// TIA Portal project "IntercambioDeDatos" (V16)

(* hardware
DEVICE "PC-System"  CPU 1515SP PC
   slot 0: "PC-System"  CPU 1515SP PC F  6ES7 677-2SBx2-0xB0  V20.8
      slot 124: "Diagbase"  Diagbase  V6.0.4
      slot 125: "PC-System"  PC Station 2.7  Station_Manager  V2.7
   slot 2: "PROFINET onboard_2"  IE General  IE_CP  V2.2.0
      slot 1: "Puerto_1"  X2 P1
   slot 3: "Software PLC_1"  CPU 1505SP F  6ES7 672-5SC11-0YA0  V2.7
      slot 3: "Display de la CPU_1"  6ES7591-1BA00-0AA0
   slot 127: "BA 2xRJ45"  BA 2xRJ45  6ES7 193-6AR00-0AA0  V0.0
      slot 32769: "Puerto_1"  X1 P1  6ES7 193-6AR00-0AA0
      slot 32770: "Puerto_2"  X1 P2  6ES7 193-6AR00-0AA0
   slot 1006: "Módulo servidor_1"  Server module  6ES7 193-6PA00-0AA0  V1.1
      slot 1: "Módulo servidor_1"  Server module
DEVICE "Dispositivo GSD_1"  GSD.Device.PN
   slot 0: "Rack"  Rack  V1.0
   slot 0: "URIODev1"  V1.0  00000
      slot 0: "V1.0"  V1.0
      slot 1: "Interface"  Interface
         slot 1: "RJ45 10/100 MBit/s"  RJ45 10/100 MBit/s
   slot 1: "1_T2O State_1"  1_T2O State  1.0
      slot 0: "1_T2O State"  1_T2O State
   slot 2: "2_T2O IO_1"  2_T2O IO  1.0
      slot 0: "2_T2O IO"  2_T2O IO
   slot 3: "3_T2O Joints_1"  3_T2O Joints  1.0
      slot 0: "3_T2O Joints"  3_T2O Joints
   slot 4: "4_T2O TCP_1"  4_T2O TCP  1.0
      slot 0: "4_T2O TCP"  4_T2O TCP
   slot 5: "5_T2O General Purpose Bit Registers_1"  5_T2O General Purpose Bit Registers  1.0
      slot 0: "5_T2O General Purpose Bit Registers"  5_T2O General Purpose Bit Registers
   slot 6: "6_T2O General Purpose Int Registers_1"  6_T2O General Purpose Int Registers  1.0
      slot 0: "6_T2O General Purpose Int Registers"  6_T2O General Purpose Int Registers
   slot 7: "7_T2O General Purpose Float Registers_1"  7_T2O General Purpose Float Registers  1.0
      slot 0: "7_T2O General Purpose Float Registers"  7_T2O General Purpose Float Registers
   slot 8: "8_O2T Robot IO_1"  8_O2T Robot IO  1.0
      slot 0: "8_O2T Robot IO"  8_O2T Robot IO
   slot 9: "9_O2T General Purpose Registers 1_1"  9_O2T General Purpose Registers 1  1.0
      slot 0: "9_O2T General Purpose Registers 1"  9_O2T General Purpose Registers 1
   slot 10: "10_O2T General Purpose Registers 2_1"  10_O2T General Purpose Registers 2  1.0
      slot 0: "10_O2T General Purpose Registers 2"  10_O2T General Purpose Registers 2
DEVICE "HMI"  KTP1200 Basic PN
   slot 0: "HMI_2"  KTP1200 Basic PN  6AV2 123-2MB03-0AX0  16.0.0.0
   slot 1: "HMI_RT_1"  KTP1200 Basic PN  6AV2 123-2MB03-0AX0  16.0.0.0
   slot 5: "HMI_2.IE_CP_1"  PROFINET Interface  16.0.0.0
      slot 1: "Interfaz PROFINET_1"  PROFINET Interface
         slot 1: "Port_1"  Port
*)

// ===== PLC "Software PLC_1"  CPU 1505SP F =====

VAR_GLOBAL   // PLC tag table "Tabla de variables estándar"
   "Flanco_Marcha" AT %M0.4 : Bool;
   "Biestable_Marcha" AT %M10.0 : Bool;
   "Tag_2" AT %M11.0 : Bool;
   "Tag_1" AT %MW20 : Int;
   "Tag_3" AT %MW22 : Int;
   "Tag_4" AT %MW24 : Int;
END_VAR

VAR_GLOBAL   // PLC tag table "IntercambioDeDatos_Variables"
   "URI" AT %I0.0 : "UR_T2O";   // Grupo de variables en donde se guardan los valores que se envian al robot
   "URO" AT %Q0.0 : "UR_O2T";   // Grupo de variables en donde se guardan los valores que llegan desde el robot
   "Marcha" AT %M0.0 : Bool;   // Variable que define en que momento debe comenzar funcionar el robot
   "Servicio_Completado" AT %M0.1 : Bool;
   "Servicio" AT %MW3 : Int;   // Variable que define el número de servicio a ejecutar
   "CantPiezas" AT %MW5 : Int;   // Variable que define la cantidad de pieza que se deben realizar.
   "Aux" AT %M1.7 : Bool;
   "No_Item_Completados" AT %MW7 : Int;
   "Item_Completado" AT %M0.2 : Bool;
   "Marcha_Reset" AT %M0.3 : Bool;
   "Flag_New_Service" AT %M0.5 : Bool;
   "MqttConnected" AT %M1.0 : Bool;
   "MqttDataReceived" AT %M1.1 : Bool;
   "Serialize" AT %M1.2 : Bool;
   "MqttSubscribed" AT %M1.3 : Bool;
   "MqttPreviousStatus" AT %MW9 : Word;
   "MqttUnsuscribed" AT %M1.4 : Bool;
   "Marcha_aux" AT %M0.6 : Bool;
   "Flanco_Service_Compl" AT %M0.7 : Bool;
   "Aux_Initial_Time_Stamp" AT %M12.0 : ULInt;
   "Aux_Final_Time_Stamp" AT %M20.0 : ULInt;
   "Aux_Service_Time_Stamp" AT %M28.0 : ULInt;
END_VAR

// folder: Common

TYPE "typeDiagnostics"
TITLE = typeDiagnostics
// Provides a structure for detailed diagnostics
   STRUCT
      status : Word;   // Status of the block or error identification when error occurred
      subfunctionStatus : DWord;   // Status or return value of called FBs, FCs and system blocks
      stateNumber : DInt;   // State in the state machine of the block where the error occurred
   END_STRUCT;
END_TYPE

// folder: LMQTT

TYPE "LMQTT_typeConnParams"
TITLE = LMQTT_typeConnParams
// Specifies connection parameters for the mqtt connection
   STRUCT
      hwId : Hw_Any;   // Hardware identifier of the interface. 0: interface is selected automatically
      connId : Conn_Ouc;   // Unique connection identifier
      brokerAddress : Struct   // Information on the MQTT broker
         qdnAddress : String;   // Fully qualified domain name of the broker. must end with a dot "."
         ipAddress : IP_V4;   // If no FQDN is used, enter ip-address of the broker instead
         port : UInt;   // Enter the port of the mqtt broker
      END_STRUCT;
      tls : Struct   // Parameters for TLS encryption
         enableTls : Bool;   // TRUE: Enables TLS, FALSE: disable TLS
         validateServerIdentity : Bool;   // TRUE: Validate server certificate, FALSE: No validation of server certificate
         brokerCert : UDInt;   // ID of the broker's certificate in TIA Portal
         clientCert : UDInt;   // ID of the client's certificate in TIA Portal
      END_STRUCT;
      keepAlive : UInt;   // Keepalive mechanism for MQTT in seconds. 0: disabled.
   END_STRUCT;
END_TYPE

// folder: LStream/DataTypes

TYPE "LStream_typeElement"
TITLE = LStream_typeElement
// describes the element for LStream libraries, by providing key-value pair and the depth of the element
   STRUCT
      "type" : SInt := -1;   // Type of element XML/JSON; -1 = inital value; 0 = Element/Object; 1 = Attribute/Array; 2 = Text/String; 3 = Number; 4 = Boolean / Type of element; -1 = inital value; 0 = Element/Object; 1 = Attribute/Array; 2 = Text
      key : String;   // Key name of element
      value : String := 'NULL';   // Value of element, null key has no value
      depth : SInt := -1;   // Depth of the key nesting
   END_STRUCT;
END_TYPE

// folder: Robot

TYPE "UR__O2T_Robot"
VERSION : 0.1
   STRUCT
      "SSM: Speed slider fraction mask" : Bool;
      Reserved_1 : Bool;
      Reserved_2 : Bool;
      Reserved_3 : Bool;
      Reserved_4 : Bool;
      Reserved_5 : Bool;
      Reserved_6 : Bool;
      Reserved_7 : Bool;
      Reserved_8_15 : USInt;
      Reserved_16_31 : UInt;
      "Speed slider fraction" : Real;
   END_STRUCT;
END_TYPE

TYPE "UR__O2T_ints"
VERSION : 0.1
   STRUCT
      Register : Array[0..11] of DInt;
   END_STRUCT;
END_TYPE

TYPE "UR__O2T_floats"
VERSION : 0.1
   STRUCT
      Register : Array[0..11] of Real;
   END_STRUCT;
END_TYPE

TYPE "UR__O2T_IOs"
VERSION : 0.1
   STRUCT
      "Standard digital output mask" : USInt;
      "Configurable digital output mask" : USInt;
      "Standard digital outputs" : USInt;
      "Configurable digital outputs" : USInt;
      "AOM: Analog output mask" : USInt;
      "AOT: Analog output types" : USInt;
      "TDOM: Tool digital output mask" : USInt;
      "TDO: Tool digital output" : USInt;
      "Standard analog output" : Array[0..1] of Real;
   END_STRUCT;
END_TYPE

TYPE "UR__O2T_bits"
VERSION : 0.1
   STRUCT
      Register : Array[0..31] of Bool;
   END_STRUCT;
END_TYPE

TYPE "UR_9_O2T_Registers"
VERSION : 0.1
   STRUCT
      Bits : "UR__O2T_bits";
      Ints : "UR__O2T_ints";
      Floats : "UR__O2T_floats";
   END_STRUCT;
END_TYPE

TYPE "UR_8_O2T_Robot_IO"
VERSION : 0.1
   STRUCT
      Robot : "UR__O2T_Robot";
      IOs : "UR__O2T_IOs";
   END_STRUCT;
END_TYPE

TYPE "UR__T2O_Safety"
VERSION : 0.1
   STRUCT
      "Safety mode" : USInt;
      Reserved_1 : USInt;
      Reserved_2 : UInt;
      "NO: Is normal mode" : Bool;
      "RD: Is reduced mode" : Bool;
      "PS: Is protective stopped" : Bool;
      "RC: Is recovery mode" : Bool;
      "SS: Is safeguard stopped" : Bool;
      "SES: Is system emergency stopped" : Bool;
      "RES: Is robot emergency stopped" : Bool;
      "ES: Is emergency stopped" : Bool;
      "VL: Is violation" : Bool;
      "FT: Is fault" : Bool;
      "ST: Is stopped due to safety" : Bool;
      Reserved_11 : Bool;
      Reserved_12 : Bool;
      Reserved_13 : Bool;
      Reserved_14 : Bool;
      Reserved_15 : Bool;
      Reserved_16_31 : UInt;
   END_STRUCT;
END_TYPE

TYPE "UR__T2O_Robot"
VERSION : 0.1
   STRUCT
      "Controller major version" : USInt;
      "Controller minor version" : USInt;
      Reserved : UInt;
      "Robot mode" : USInt;
      "Real time machine seconds" : USInt;
      "Real time machine milliseconds" : UInt;
      "Real time machine minutes" : USInt;
      "Real time machine hours" : USInt;
      "Real time machine days" : UInt;
      "Robot current [A]" : Real;
      "PW: Is power on" : Bool;
      "PR: Is program running" : Bool;
      "TB: Is teach button pressed" : Bool;
      "PB: Is power button pressed" : Bool;
      Reserved_4 : Bool;
      Reserved_5 : Bool;
      Reserved_6 : Bool;
      Reserved_7 : Bool;
      Reserved_8_15 : USInt;
      Reserved_16_31 : UInt;
      "Speed slider fraction" : Real;
   END_STRUCT;
END_TYPE

TYPE "UR__T2O_Tool"
VERSION : 0.1
   STRUCT
      "Tool mode" : USInt;
      Reserved_7_15 : USInt;
      Reserved_16_31 : UInt;
      "TDI: Tool Digital Inputs" : USInt;
      "TDO: Tool Digital Outputs" : USInt;
      "TAIT: Tool Analog Input Types" : USInt;
      Reserved_24_31 : USInt;
      "Tool analog input [A or V]" : Array[0..1] of Real;
      "Tool output voltage [V]" : Real;
      "Tool current [A]" : Real;
   END_STRUCT;
END_TYPE

TYPE "UR_O2T"
VERSION : 0.1
   STRUCT
      "Robot IO" : "UR_8_O2T_Robot_IO";
      "Reg 1" : "UR_9_O2T_Registers";
      "Reg 2" : "UR_9_O2T_Registers";
   END_STRUCT;
END_TYPE

TYPE "UR_4_T2O_TCP"
VERSION : 0.1
   STRUCT
      "TCP Position (X,Y,Z) [m]" : Array[0..2] of Real;
      "TCP Position (RX,RY,RZ) [rad]" : Array[0..2] of Real;
      "TCP velocity (X,Y,Z) [m/s]" : Array[0..2] of Real;
      "TCP velocity (RX,RY,RZ) [rad/s]" : Array[0..2] of Real;
      "TCP force (X,Y,Z) [N]" : Array[0..2] of Real;
      "TCP torque (X,Y,Z) [Nm]" : Array[0..2] of Real;
      "TCP force scalar [N]" : Real;
   END_STRUCT;
END_TYPE

TYPE "UR_3_T2O_Joints"
VERSION : 0.1
   STRUCT
      "Joint position [rad]" : Array[0..5] of Real;
      "Joint velocity [rad/s]" : Array[0..5] of Real;
      "Joint current [A]" : Array[0..5] of Real;
      "Joint temperature [°C]" : Array[0..5] of Real;
      "Joint mode" : Array[0..5] of USInt;
      Reserved_9 : UInt;
   END_STRUCT;
END_TYPE

TYPE "UR_2_T2O_IO"
VERSION : 0.1
   STRUCT
      IOs : "UR__T2O_IOs";
      Tool : "UR__T2O_Tool";
   END_STRUCT;
END_TYPE

TYPE "UR_1_T2O_State"
VERSION : 0.1
   STRUCT
      Robot : "UR__T2O_Robot";
      Safety : "UR__T2O_Safety";
   END_STRUCT;
END_TYPE

TYPE "UR_7_T2O_FloatRegisters"
VERSION : 0.1
   STRUCT
      Register : Array[0..23] of Real;
   END_STRUCT;
END_TYPE

TYPE "UR_6_T2O_IntRegisters"
VERSION : 0.1
   STRUCT
      Register : Array[0..23] of DInt;
   END_STRUCT;
END_TYPE

TYPE "UR_T2O"
VERSION : 0.1
   STRUCT
      State : "UR_1_T2O_State";
      IO : "UR_2_T2O_IO";
      Joints : "UR_3_T2O_Joints";
      TCP : "UR_4_T2O_TCP";
      Bits : "UR_5_T2O_BitRegisters";
      Ints : "UR_6_T2O_IntRegisters";
      Floats : "UR_7_T2O_FloatRegisters";
   END_STRUCT;
END_TYPE

TYPE "UR__T2O_IOs"
VERSION : 0.1
   STRUCT
      "Standard digital inputs" : USInt;
      "Configurable digital inputs" : USInt;
      "Standard digital outputs" : USInt;
      "Configurable digital outputs" : USInt;
      "Analog I/O types" : USInt;
      Reserved_8_15 : USInt;
      Reserved_16_31 : UInt;
      "Standard analog input [A or V]" : Array[0..1] of Real;
      "Standard analog output [A or V]" : Array[0..1] of Real;
      "I/O current [A]" : Real;
      "Euromap67 input bits" : Array[0..31] of Bool;
      "Euromap67 output bits" : Array[0..31] of Bool;
      "Euromap67 24V voltage" : Real;
      "Euromap67 24V current" : Real;
   END_STRUCT;
END_TYPE

TYPE "UR_5_T2O_BitRegisters"
VERSION : 0.1
   STRUCT
      Register : Array[0..63] of Bool;
   END_STRUCT;
END_TYPE

// folder: (top level)

DATA_BLOCK "Main_Safety_RTG1_DB"   // DB1, F_DB
{ S7_Optimized_Access := 'TRUE' }
NAME : FUSI
VERSION : 0.1
// stored: InstanceOfName Main_Safety_RTG1
"Main_Safety_RTG1"
BEGIN
END_DATA_BLOCK

DATA_BLOCK "MqttDB"   // DB3
{ S7_Optimized_Access := 'TRUE' }
AUTHOR : Siemens
FAMILY : LMQTT
VERSION : 1.0
   VAR
      control : Struct
         connect : Bool;
         publish : Bool;
         subscribe : Bool;
         unsubscribe : Bool;
      END_STRUCT;
      output : Struct
         valid : Bool;
         done : Bool;
         busy : Bool;
         error : Bool;
         status : Word;
         diagnostics : "typeDiagnostics";
      END_STRUCT;
      connparams : "LMQTT_typeConnParams";
      clientid : WString[20] := WSTRING#'Alazne';
      username : WString[20];
      password : WString[20];
      willtopic : WString[20] := WSTRING#'willTopic';
      willMessage : Array[0..99] of Byte;
      willmesscnt : UInt := 10;
      qos : USInt := 0;
      topic : WString[100] := WSTRING#'Operation';
      message : Array[0..999] of Byte;
      pubMessageCnt : UDInt := 1;
      retain : Bool;
      receivedTopic : WString[200];
      receivedmessage : Array[0..999] of Byte;
      receivedMsgLen : UDInt;
      receivedMsgStatus : USInt;
      dadoRecebido : String[100];
      dadoEnviado : String[100];
   END_VAR
BEGIN
   connparams.connId := 16#0001;
   connparams.brokerAddress.port := 1883;
   willMessage[0] := 16#6F;
   willMessage[1] := 16#66;
   willMessage[2] := 16#66;
   willMessage[3] := 16#6C;
   willMessage[4] := 16#69;
   willMessage[5] := 16#6E;
   willMessage[6] := 16#65;
   message[0] := 53;
   connparams.brokerAddress.ipAddress.ADDR[1] := 192;
   connparams.brokerAddress.ipAddress.ADDR[2] := 168;
   connparams.brokerAddress.ipAddress.ADDR[3] := 2;
   connparams.brokerAddress.ipAddress.ADDR[4] := 151;
   connparams.keepAlive := 30;   // Periodo de tiempo durante el cual se considera que una conexión esta viva sin que hay consexión entre el cliente y el bróker.
   connparams.hwId := 0;
END_DATA_BLOCK

DATA_BLOCK "AASassetDB"   // DB5
{ S7_Optimized_Access := 'TRUE' }
VERSION : 0.1
   VAR
      Control : Struct
         Flag_New_Service : Bool;
         Flag_Item_Completed : Bool;
         Flag_Service_Completed : Bool;
      END_STRUCT;
      Agent2PLC : Struct
         Id : Struct
            Machine_Reference : UDInt;
            Order_Reference : UDInt;
            Batch_Reference : UDInt;
            Ref_Subproduct_Type : UDInt;
         END_STRUCT;
         Operation : Struct
            Ref_Service_Type : UDInt;
            No_of_Items : USInt;
         END_STRUCT;
      END_STRUCT;
      PLC2Agent : Struct
         Id : Struct
            Machine_Reference : UDInt;
            Order_Reference : UDInt;
            Batch_Reference : UDInt;
            Ref_Subproduct_Type : UDInt;
            Ref_Service_Type : UDInt;
            Item_Number : USInt;
         END_STRUCT;
         Data : Struct
            Initial_Time_Stamp : LDT;
            Final_Time_Stamp : LDT;
            Service_Time_Stamp : LDT;
         END_STRUCT;
      END_STRUCT;
   END_VAR
BEGIN
END_DATA_BLOCK

DATA_BLOCK "JSON_DeserializParamDB"   // DB9
{ S7_Optimized_Access := 'TRUE' }
VERSION : 0.1
   VAR
      execute : Bool;
      search : Bool;
      jsonByteArray : Array[0..999] of Byte;
      tree : Array[0..999] of "LStream_typeElement";
      resultCount : Int;
      out : Struct
         done : Bool;
         busy : Bool;
         error : Bool;
         status : Word;
         resultCount : Int;
      END_STRUCT;
   END_VAR
BEGIN
END_DATA_BLOCK

DATA_BLOCK "JSON_SerializParamDB"   // DB10
{ S7_Optimized_Access := 'TRUE' }
VERSION : 0.1
   VAR
      execute : Bool;
      out : Struct
         done : Bool;
         busy : Bool;
         error : Bool;
         status : Word;
      END_STRUCT;
      tree : Array[0..999] of "LStream_typeElement";
      jsonByteArray : Array[0..999] of Byte;
      resultCount : Int;
   END_VAR
BEGIN
   tree[0]."type" := 0;
   tree[0].key := 'Control';
   tree[0].depth := 0;
   tree[1]."type" := 4;
   tree[1].key := 'Flag_Item_Completed';
   tree[1].depth := 1;
   tree[2]."type" := 4;
   tree[2].key := 'Flag_Service_Completed';
   tree[2].depth := 1;
   tree[3]."type" := 0;
   tree[3].key := 'Id';
   tree[3].depth := 0;
   tree[4]."type" := 3;
   tree[4].key := 'Machine_Reference';
   tree[4].depth := 1;
   tree[5]."type" := 3;
   tree[5].key := 'Order_Reference';
   tree[5].depth := 1;
   tree[6]."type" := 3;
   tree[6].key := 'Batch_Reference';
   tree[6].depth := 1;
   tree[7]."type" := 3;
   tree[7].key := 'Ref_Subproduct_Type';
   tree[7].depth := 1;
   tree[8].key := 'Ref_Service_Type';
   tree[8]."type" := 3;
   tree[8].depth := 1;
   tree[9]."type" := 3;
   tree[9].key := 'Item_Number';
   tree[9].depth := 1;
   tree[10]."type" := 0;
   tree[10].key := 'Data';
   tree[10].depth := 0;
   tree[11]."type" := 3;
   tree[11].key := 'Initial_Time_Stamp';
   tree[11].depth := 1;
   tree[12]."type" := 3;
   tree[12].key := 'Final_Time_Stamp';
   tree[12].depth := 1;
   tree[13]."type" := 3;
   tree[13].key := 'Service_Time_Stamp';
   tree[13].depth := 1;
END_DATA_BLOCK

// folder: LMQTT

DATA_BLOCK "LMQTT_Client_DB"   // DB2
{ S7_Optimized_Access := 'TRUE' }
AUTHOR : SUP
FAMILY : LMQTT
VERSION : 3.0
// stored: InstanceOfName LMQTT_Client
"LMQTT_Client"
BEGIN
END_DATA_BLOCK

// folder: LStream

DATA_BLOCK "LStream_JsonDeserializer_DB"   // DB7
{ S7_Optimized_Access := 'TRUE' }
AUTHOR : DI_FA_S_SUP_EuC
FAMILY : LStream
VERSION : 1.0
// stored: InstanceOfName LStream_JsonDeserializer
"LStream_JsonDeserializer"
BEGIN
END_DATA_BLOCK

DATA_BLOCK "LStream_JsonSerializer_DB"   // DB8
{ S7_Optimized_Access := 'TRUE' }
AUTHOR : DI_FA_S_SUP_EuC
FAMILY : LStream
VERSION : 1.0
// stored: InstanceOfName LStream_JsonSerializer
"LStream_JsonSerializer"
BEGIN
END_DATA_BLOCK

// folder: (top level)

FUNCTION_BLOCK "Main_Safety_RTG1"   // FB1, F_FBD
{ S7_Optimized_Access := 'TRUE' }
BEGIN
END_FUNCTION_BLOCK

FUNCTION "Outputs2LStreamTree" : Void   // FC1, SCL
{ S7_Optimized_Access := 'TRUE' }
VERSION : 0.1
BEGIN
   // Asignación de valores 
   (* "JSON_SerializParamDB".tree[1].value := "AASassetDb".Control.Flag_Item_Completed; *)

   (* "JSON_SerializParamDB".tree[1].value := 'false';
   "JSON_SerializParamDB".tree[2].value := 'false'; *)
   (* "JSON_SerializParamDB".tree[4].value := '123';
   "JSON_SerializParamDB".tree[5].value := '22';
   "JSON_SerializParamDB".tree[6].value := '33';
   "JSON_SerializParamDB".tree[7].value := '99'; *)

   IF "AASassetDB".Control.Flag_Service_Completed = 1 THEN
       "JSON_SerializParamDB".tree[2].value := 'true';
   ELSE
       "JSON_SerializParamDB".tree[2].value := 'false';
   END_IF;

   IF "AASassetDB".Control.Flag_Item_Completed = 1 THEN
       "JSON_SerializParamDB".tree[1].value := 'true';
   ELSE
       "JSON_SerializParamDB".tree[1].value := 'false';
   END_IF;

   "JSON_SerializParamDB".tree[4].value := UDINT_TO_STRING("AASassetDB".PLC2Agent.Id.Machine_Reference);
   "JSON_SerializParamDB".tree[5].value := UDINT_TO_STRING("AASassetDB".PLC2Agent.Id.Order_Reference);
   "JSON_SerializParamDB".tree[6].value := UDINT_TO_STRING("AASassetDB".PLC2Agent.Id.Batch_Reference);
   "JSON_SerializParamDB".tree[7].value := UDINT_TO_STRING("AASassetDB".PLC2Agent.Id.Ref_Subproduct_Type);
   "JSON_SerializParamDB".tree[8].value := UDINT_TO_STRING("AASassetDB".PLC2Agent.Id.Ref_Service_Type);
   "JSON_SerializParamDB".tree[9].value := USINT_TO_STRING("AASassetDB".PLC2Agent.Id.Item_Number);

   "JSON_SerializParamDB".tree[11].value := ULINT_TO_STRING(LDT_TO_ULINT("AASassetDB".PLC2Agent.Data.Initial_Time_Stamp));
   "JSON_SerializParamDB".tree[12].value := ULINT_TO_STRING(LDT_TO_ULINT("AASassetDB".PLC2Agent.Data.Final_Time_Stamp));
   "JSON_SerializParamDB".tree[13].value := ULINT_TO_STRING(LDT_TO_ULINT("AASassetDB".PLC2Agent.Data.Service_Time_Stamp));
END_FUNCTION

FUNCTION "LStreamTree2Inputs" : Void   // FC3, SCL
{ S7_Optimized_Access := 'TRUE' }
VERSION : 0.1
   VAR_TEMP
      Indice : Int;
   END_VAR
BEGIN
   // Volcado de los valores recibidos del bróker en las variables del DB.

   // Id
   "AASassetDB".Agent2PLC.Id.Machine_Reference := STRING_TO_UDINT("JSON_DeserializParamDB".tree[8].value);
   "AASassetDB".Agent2PLC.Id.Order_Reference := STRING_TO_UDINT("JSON_DeserializParamDB".tree[7].value);
   "AASassetDB".Agent2PLC.Id.Batch_Reference := STRING_TO_UDINT("JSON_DeserializParamDB".tree[5].value);
   "AASassetDB".Agent2PLC.Id.Ref_Subproduct_Type := STRING_TO_UDINT("JSON_DeserializParamDB".tree[6].value);

   // Operation
   "AASassetDB".Agent2PLC.Operation.Ref_Service_Type := STRING_TO_UDINT("JSON_DeserializParamDB".tree[11].value);
   "AASassetDB".Agent2PLC.Operation.No_of_Items := STRING_TO_USINT("JSON_DeserializParamDB".tree[10].value);
END_FUNCTION

ORGANIZATION_BLOCK "Main"   // OB1, LAD, ProgramCycle
TITLE = "Main Program Sweep (Cycle)"
{ S7_Optimized_Access := 'TRUE' }
VERSION : 0.1
   VAR_INPUT
      Initial_Call : Bool;   // Initial call of this OB
      Remanence : Bool;   // =True, if remanent data are available
   END_VAR
   VAR_TEMP
      FlancoNeg_Item_Completed : Bool;
      FlancoPos_Item_Completed : Bool;
   END_VAR
   VAR_TEMP   // added for the SCL form of the ladder/FBD networks
      _w1 : Bool;
      _w2 : Bool;
   END_VAR
BEGIN

REGION Network 1: Cliente MQTT
   // En este segmento nos encargamos tanto de la suscripción a un tópico como de las publicaciones que se realizarán en el tópico de publicaciones.
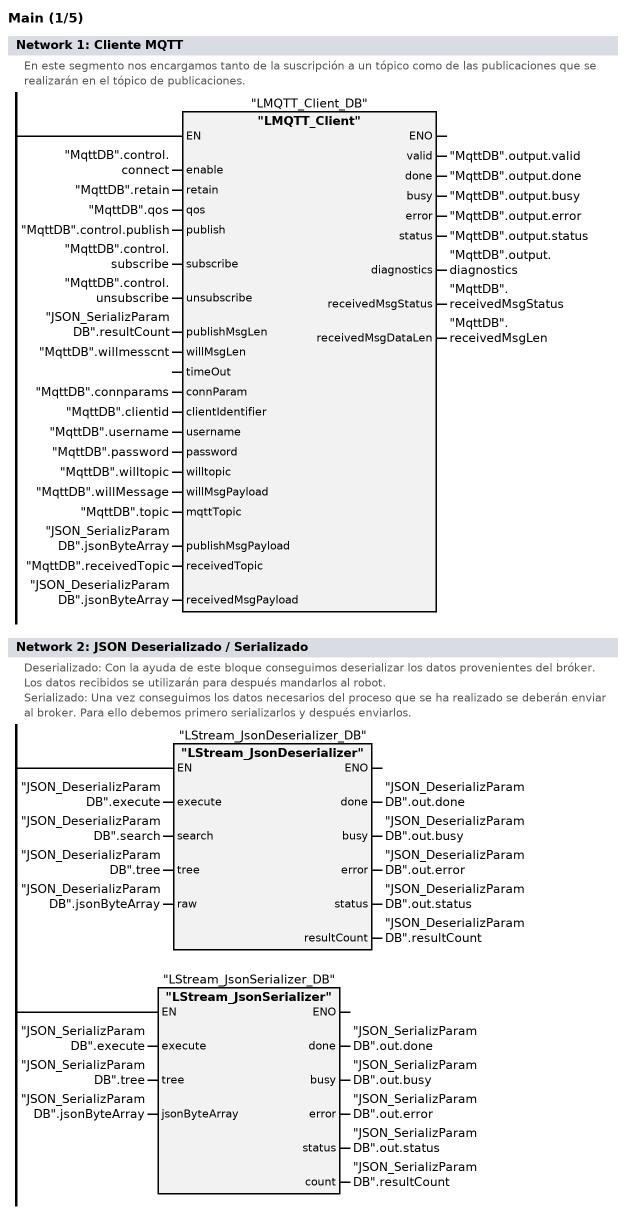
   RUNG wire#powerrail
      "LMQTT_Client_DB"(enable := "MqttDB".control.connect, retain := "MqttDB".retain, qos := "MqttDB".qos, publish := "MqttDB".control.publish, subscribe := "MqttDB".control.subscribe, unsubscribe := "MqttDB".control.unsubscribe, publishMsgLen := "JSON_SerializParamDB".resultCount, willMsgLen := "MqttDB".willmesscnt, timeOut :=, connParam := "MqttDB".connparams, clientIdentifier := "MqttDB".clientid, username := "MqttDB".username, password := "MqttDB".password, willtopic := "MqttDB".willtopic, willMsgPayload := "MqttDB".willMessage, mqttTopic := "MqttDB".topic, publishMsgPayload := "JSON_SerializParamDB".jsonByteArray, receivedTopic := "MqttDB".receivedTopic, receivedMsgPayload := "JSON_DeserializParamDB".jsonByteArray, valid => "MqttDB".output.valid, done => "MqttDB".output.done, busy => "MqttDB".output.busy, error => "MqttDB".output.error, status => "MqttDB".output.status, diagnostics => "MqttDB".output.diagnostics, receivedMsgStatus => "MqttDB".receivedMsgStatus, receivedMsgDataLen => "MqttDB".receivedMsgLen)
   END_RUNG
   // the same network as SCL:
   "LMQTT_Client_DB"(enable := "MqttDB".control.connect,   // "LMQTT_Client"
                     retain := "MqttDB".retain,
                     qos := "MqttDB".qos,
                     publish := "MqttDB".control.publish,
                     subscribe := "MqttDB".control.subscribe,
                     unsubscribe := "MqttDB".control.unsubscribe,
                     publishMsgLen := "JSON_SerializParamDB".resultCount,
                     willMsgLen := "MqttDB".willmesscnt,
                     connParam := "MqttDB".connparams,
                     clientIdentifier := "MqttDB".clientid,
                     username := "MqttDB".username,
                     password := "MqttDB".password,
                     willtopic := "MqttDB".willtopic,
                     willMsgPayload := "MqttDB".willMessage,
                     mqttTopic := "MqttDB".topic,
                     publishMsgPayload := "JSON_SerializParamDB".jsonByteArray,
                     receivedTopic := "MqttDB".receivedTopic,
                     receivedMsgPayload := "JSON_DeserializParamDB".jsonByteArray,
                     valid => "MqttDB".output.valid,
                     done => "MqttDB".output.done,
                     busy => "MqttDB".output.busy,
                     error => "MqttDB".output.error,
                     status => "MqttDB".output.status,
                     diagnostics => "MqttDB".output.diagnostics,
                     receivedMsgStatus => "MqttDB".receivedMsgStatus,
                     receivedMsgDataLen => "MqttDB".receivedMsgLen);
END_REGION

REGION Network 2: JSON Deserializado / Serializado
   // Deserializado: Con la ayuda de este bloque conseguimos deserializar los datos provenientes del bróker. 
   // Los datos recibidos se utilizarán para después mandarlos al robot.
   // 
   // Serializado: Una vez conseguimos los datos necesarios del proceso que se ha realizado se deberán enviar al broker. Para ello debemos primero serializarlos y después enviarlos.
   RUNG wire#powerrail
      "LStream_JsonDeserializer_DB"(execute := "JSON_DeserializParamDB".execute, search := "JSON_DeserializParamDB".search, tree := "JSON_DeserializParamDB".tree, raw := "JSON_DeserializParamDB".jsonByteArray, done => "JSON_DeserializParamDB".out.done, busy => "JSON_DeserializParamDB".out.busy, error => "JSON_DeserializParamDB".out.error, status => "JSON_DeserializParamDB".out.status, resultCount => "JSON_DeserializParamDB".resultCount)
   END_RUNG
   RUNG wire#powerrail
      "LStream_JsonSerializer_DB"(execute := "JSON_SerializParamDB".execute, tree := "JSON_SerializParamDB".tree, jsonByteArray := "JSON_SerializParamDB".jsonByteArray, done => "JSON_SerializParamDB".out.done, busy => "JSON_SerializParamDB".out.busy, error => "JSON_SerializParamDB".out.error, status => "JSON_SerializParamDB".out.status, count => "JSON_SerializParamDB".resultCount)
   END_RUNG
   // the same network as SCL:
   "LStream_JsonDeserializer_DB"(execute := "JSON_DeserializParamDB".execute,   // "LStream_JsonDeserializer"
                           search := "JSON_DeserializParamDB".search,
                           tree := "JSON_DeserializParamDB".tree,
                           raw := "JSON_DeserializParamDB".jsonByteArray,
                           done => "JSON_DeserializParamDB".out.done,
                           busy => "JSON_DeserializParamDB".out.busy,
                           error => "JSON_DeserializParamDB".out.error,
                           status => "JSON_DeserializParamDB".out.status,
                           resultCount => "JSON_DeserializParamDB".resultCount);
   "LStream_JsonSerializer_DB"(execute := "JSON_SerializParamDB".execute,   // "LStream_JsonSerializer"
                           tree := "JSON_SerializParamDB".tree,
                           jsonByteArray := "JSON_SerializParamDB".jsonByteArray,
                           done => "JSON_SerializParamDB".out.done,
                           busy => "JSON_SerializParamDB".out.busy,
                           error => "JSON_SerializParamDB".out.error,
                           status => "JSON_SerializParamDB".out.status,
                           count => "JSON_SerializParamDB".resultCount);
END_REGION

REGION Network 3: Asignación de valores dependiendo del valor de STATUS.
   // En el momento que el valor de MqttDB sea igual a 16#7000 significa que no hay ningún tipo de conexión por lo que a los valores se les asigna un RESET.
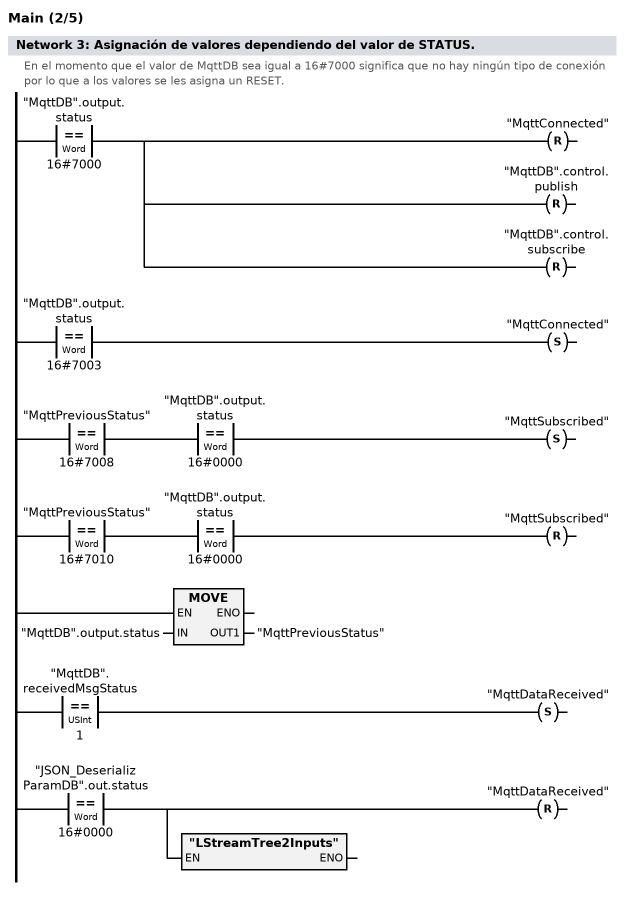
   RUNG wire#powerrail
      { S7_Templates := "SrcType := Word" } EQ_Contact(in1 := "MqttDB".output.status, in2 := 16#7000)
      wire#w1
      R_Coil( "MqttConnected" )
   END_RUNG
   RUNG wire#w1
      R_Coil( "MqttDB".control.publish )
   END_RUNG
   RUNG wire#w1
      R_Coil( "MqttDB".control.subscribe )
   END_RUNG
   RUNG wire#powerrail
      { S7_Templates := "SrcType := Word" } EQ_Contact(in1 := "MqttDB".output.status, in2 := 16#7003)
      S_Coil( "MqttConnected" )
   END_RUNG
   RUNG wire#powerrail
      { S7_Templates := "SrcType := Word" } EQ_Contact(in1 := "MqttPreviousStatus", in2 := 16#7008)
      { S7_Templates := "SrcType := Word" } EQ_Contact(in1 := "MqttDB".output.status, in2 := 16#0000)
      S_Coil( "MqttSubscribed" )
   END_RUNG
   RUNG wire#powerrail
      { S7_Templates := "SrcType := Word" } EQ_Contact(in1 := "MqttPreviousStatus", in2 := 16#7010)
      { S7_Templates := "SrcType := Word" } EQ_Contact(in1 := "MqttDB".output.status, in2 := 16#0000)
      R_Coil( "MqttSubscribed" )
   END_RUNG
   RUNG wire#powerrail
      Move(in := "MqttDB".output.status, out1 => "MqttPreviousStatus")
   END_RUNG
   RUNG wire#powerrail
      { S7_Templates := "SrcType := USInt" } EQ_Contact(in1 := "MqttDB".receivedMsgStatus, in2 := 1)
      S_Coil( "MqttDataReceived" )
   END_RUNG
   RUNG wire#powerrail
      { S7_Templates := "SrcType := Word" } EQ_Contact(in1 := "JSON_DeserializParamDB".out.status, in2 := 16#0000)
      wire#w2
      R_Coil( "MqttDataReceived" )
   END_RUNG
   RUNG wire#w2
      "LStreamTree2Inputs"()
   END_RUNG
   // the same network as SCL:
   IF "MqttDB".output.status = 16#7000 THEN
       "MqttConnected" := FALSE;
       "MqttDB".control.publish := FALSE;
       "MqttDB".control.subscribe := FALSE;
   END_IF;
   IF "MqttDB".output.status = 16#7003 THEN "MqttConnected" := TRUE; END_IF;
   IF ("MqttPreviousStatus" = 16#7008) AND ("MqttDB".output.status = 16#0000) THEN
       "MqttSubscribed" := TRUE;
   END_IF;
   IF ("MqttPreviousStatus" = 16#7010) AND ("MqttDB".output.status = 16#0000) THEN
       "MqttSubscribed" := FALSE;
   END_IF;
   "MqttPreviousStatus" := "MqttDB".output.status;
   IF "MqttDB".receivedMsgStatus = 1 THEN "MqttDataReceived" := TRUE; END_IF;
   IF "JSON_DeserializParamDB".out.status = 16#0000 THEN
       "MqttDataReceived" := FALSE;
       "LStreamTree2Inputs"();
   END_IF;
END_REGION

REGION Network 4: Marcha y Operacion Finalizada
   // Flag_New_Service -> esta variable se pone en TRUE en el momento que queramos comenzar con un nuevo servicio. llega desde el agente
   // 
   // Flag_Service_Completed -> Indicador que define que el servicio a realizar se ha finalizado. Se define en el robot y se manda al agente.
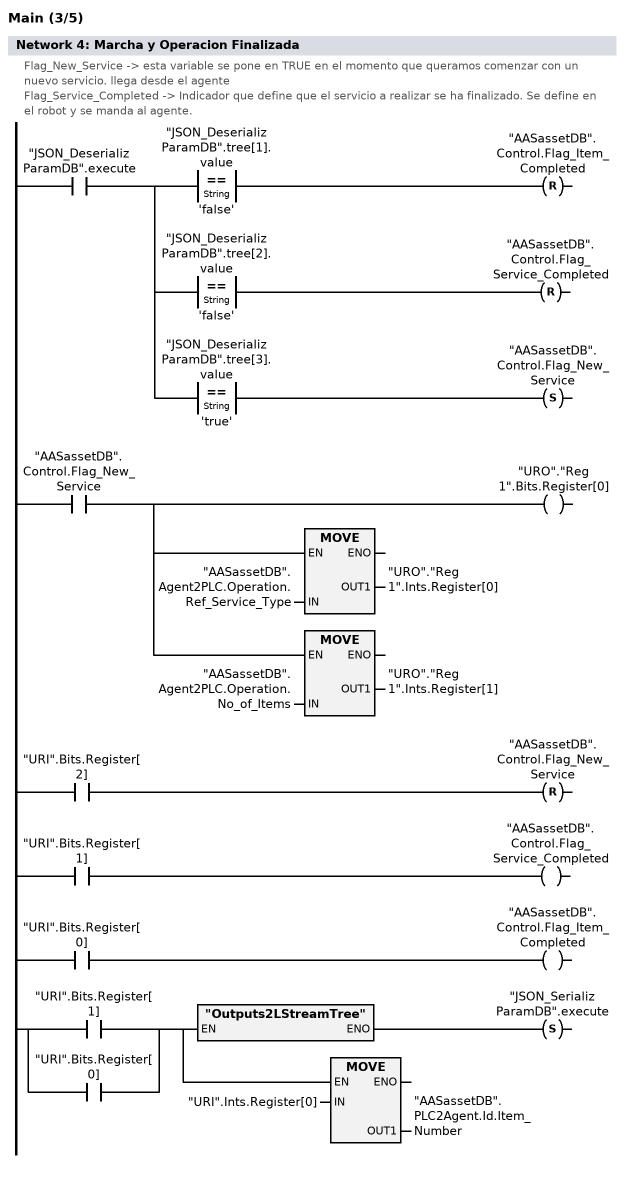
   RUNG wire#powerrail
      Contact( "JSON_DeserializParamDB".execute )
      wire#w1
      { S7_Templates := "SrcType := String" } EQ_Contact(in1 := "JSON_DeserializParamDB".tree[1].value, in2 := 'false')
      R_Coil( "AASassetDB".Control.Flag_Item_Completed )
   END_RUNG
   RUNG wire#w1
      { S7_Templates := "SrcType := String" } EQ_Contact(in1 := "JSON_DeserializParamDB".tree[2].value, in2 := 'false')
      R_Coil( "AASassetDB".Control.Flag_Service_Completed )
   END_RUNG
   RUNG wire#w1
      { S7_Templates := "SrcType := String" } EQ_Contact(in1 := "JSON_DeserializParamDB".tree[3].value, in2 := 'true')
      S_Coil( "AASassetDB".Control.Flag_New_Service )
   END_RUNG
   RUNG wire#powerrail
      Contact( "AASassetDB".Control.Flag_New_Service )
      wire#w2
      Coil( "URO"."Reg 1".Bits.Register[0] )
   END_RUNG
   RUNG wire#w2
      Move(in := "AASassetDB".Agent2PLC.Operation.Ref_Service_Type, out1 => "URO"."Reg 1".Ints.Register[0])
   END_RUNG
   RUNG wire#w2
      Move(in := "AASassetDB".Agent2PLC.Operation.No_of_Items, out1 => "URO"."Reg 1".Ints.Register[1])
   END_RUNG
   RUNG wire#powerrail
      Contact( "URI".Bits.Register[2] )
      R_Coil( "AASassetDB".Control.Flag_New_Service )
   END_RUNG
   RUNG wire#powerrail
      Contact( "URI".Bits.Register[1] )
      Coil( "AASassetDB".Control.Flag_Service_Completed )
   END_RUNG
   RUNG wire#powerrail
      Contact( "URI".Bits.Register[0] )
      Coil( "AASassetDB".Control.Flag_Item_Completed )
   END_RUNG
   RUNG wire#powerrail
      Contact( "URI".Bits.Register[1] )
      wire#w3
      "Outputs2LStreamTree"()
      S_Coil( "JSON_SerializParamDB".execute )
   END_RUNG
   RUNG wire#powerrail
      Contact( "URI".Bits.Register[0] )
   END_RUNG wire#w3
   RUNG wire#w3
      Move(in := "URI".Ints.Register[0], out1 => "AASassetDB".PLC2Agent.Id.Item_Number)
   END_RUNG
   // the same network as SCL:
   IF "JSON_DeserializParamDB".execute AND ("JSON_DeserializParamDB".tree[1].value = 'false') THEN
       "AASassetDB".Control.Flag_Item_Completed := FALSE;
   END_IF;
   IF "JSON_DeserializParamDB".execute AND ("JSON_DeserializParamDB".tree[2].value = 'false') THEN
       "AASassetDB".Control.Flag_Service_Completed := FALSE;
   END_IF;
   IF "JSON_DeserializParamDB".execute AND ("JSON_DeserializParamDB".tree[3].value = 'true') THEN
       "AASassetDB".Control.Flag_New_Service := TRUE;
   END_IF;
   "URO"."Reg 1".Bits.Register[0] := "AASassetDB".Control.Flag_New_Service;
   IF "AASassetDB".Control.Flag_New_Service THEN
       "URO"."Reg 1".Ints.Register[0] := "AASassetDB".Agent2PLC.Operation.Ref_Service_Type;
       "URO"."Reg 1".Ints.Register[1] := "AASassetDB".Agent2PLC.Operation.No_of_Items;
   END_IF;
   IF "URI".Bits.Register[2] THEN "AASassetDB".Control.Flag_New_Service := FALSE; END_IF;
   "AASassetDB".Control.Flag_Service_Completed := "URI".Bits.Register[1];
   "AASassetDB".Control.Flag_Item_Completed := "URI".Bits.Register[0];
   #_w2 := "URI".Bits.Register[1] OR "URI".Bits.Register[0];
   "Outputs2LStreamTree"(EN := "URI".Bits.Register[1] OR "URI".Bits.Register[0], ENO => #_w1);
   IF #_w1 THEN "JSON_SerializParamDB".execute := TRUE; END_IF;
   IF #_w2 THEN "AASassetDB".PLC2Agent.Id.Item_Number := "URI".Ints.Register[0]; END_IF;
END_REGION

REGION Network 5: Tópicos
   // En este segmento se definen los dos tópicos con los que vamos a trabajar. 
   // Un tópico será para publicar y el otra se utiliza en la suscripción.
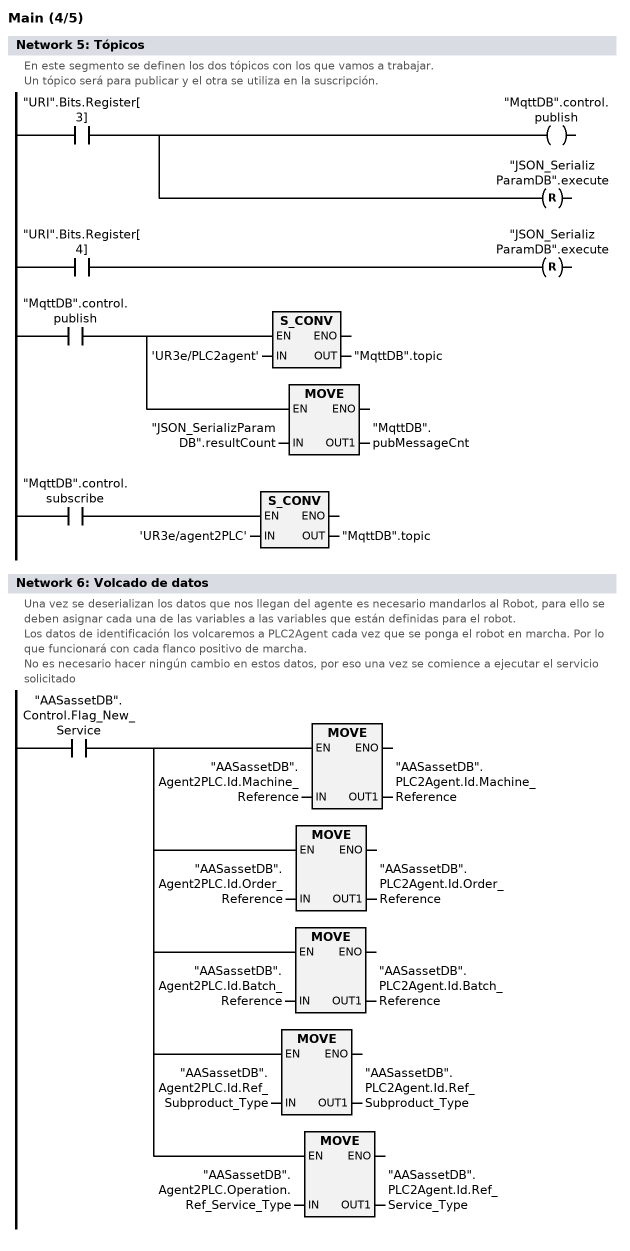
   "MqttDB".control.publish := "URI".Bits.Register[3];
   IF "URI".Bits.Register[3] THEN "JSON_SerializParamDB".execute := FALSE; END_IF;
   IF "URI".Bits.Register[4] THEN "JSON_SerializParamDB".execute := FALSE; END_IF;
   #_w1 := "MqttDB".control.publish;
   IF #_w1 THEN
       "MqttDB".topic := S_CONV(IN := 'UR3e/PLC2agent');
       "MqttDB".pubMessageCnt := "JSON_SerializParamDB".resultCount;
   END_IF;
   IF "MqttDB".control.subscribe THEN "MqttDB".topic := S_CONV(IN := 'UR3e/agent2PLC'); END_IF;
END_REGION

REGION Network 6: Volcado de datos
   // Una vez se deserializan los datos que nos llegan del agente es necesario mandarlos al Robot, para ello se deben asignar cada una de las variables a las variables que están definidas para el robot.
   // Los datos de identificación los volcaremos a PLC2Agent cada vez que se ponga el robot en marcha. Por lo que funcionará con cada flanco positivo de marcha.
   // 
   // No es necesario hacer ningún cambio en estos datos, por eso una vez se comience a ejecutar el servicio solicitado
   RUNG wire#powerrail
      Contact( "AASassetDB".Control.Flag_New_Service )
      wire#w1
      Move(in := "AASassetDB".Agent2PLC.Id.Machine_Reference, out1 => "AASassetDB".PLC2Agent.Id.Machine_Reference)
   END_RUNG
   RUNG wire#w1
      Move(in := "AASassetDB".Agent2PLC.Id.Order_Reference, out1 => "AASassetDB".PLC2Agent.Id.Order_Reference)
   END_RUNG
   RUNG wire#w1
      Move(in := "AASassetDB".Agent2PLC.Id.Batch_Reference, out1 => "AASassetDB".PLC2Agent.Id.Batch_Reference)
   END_RUNG
   RUNG wire#w1
      Move(in := "AASassetDB".Agent2PLC.Id.Ref_Subproduct_Type, out1 => "AASassetDB".PLC2Agent.Id.Ref_Subproduct_Type)
   END_RUNG
   RUNG wire#w1
      Move(in := "AASassetDB".Agent2PLC.Operation.Ref_Service_Type, out1 => "AASassetDB".PLC2Agent.Id.Ref_Service_Type)
   END_RUNG
   // the same network as SCL:
   IF "AASassetDB".Control.Flag_New_Service THEN
       "AASassetDB".PLC2Agent.Id.Machine_Reference := "AASassetDB".Agent2PLC.Id.Machine_Reference;
       "AASassetDB".PLC2Agent.Id.Order_Reference := "AASassetDB".Agent2PLC.Id.Order_Reference;
       "AASassetDB".PLC2Agent.Id.Batch_Reference := "AASassetDB".Agent2PLC.Id.Batch_Reference;
       "AASassetDB".PLC2Agent.Id.Ref_Subproduct_Type := "AASassetDB".Agent2PLC.Id.Ref_Subproduct_Type;
       "AASassetDB".PLC2Agent.Id.Ref_Service_Type := "AASassetDB".Agent2PLC.Operation.Ref_Service_Type;
   END_IF;
END_REGION

REGION Network 7: Time Stamp
   // En este segmento se definen las variables que definen la hora y el dia en el que se realiza el servicio solicitado.
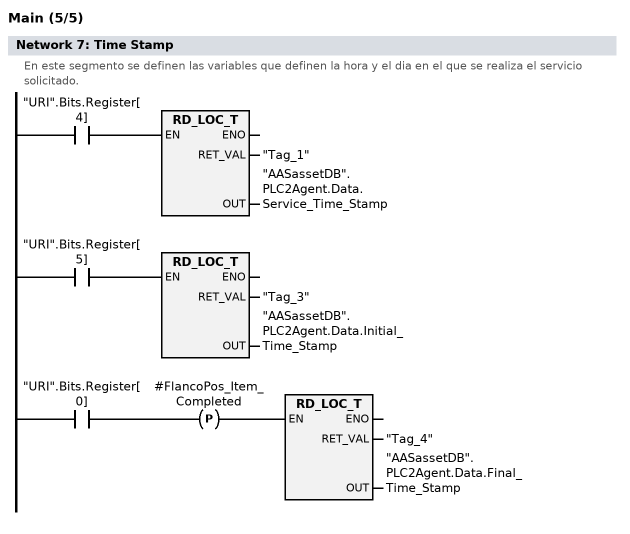
   IF "URI".Bits.Register[4] THEN
       "Tag_1" := RD_LOC_T(OUT => "AASassetDB".PLC2Agent.Data.Service_Time_Stamp);
   END_IF;
   IF "URI".Bits.Register[5] THEN
       "Tag_3" := RD_LOC_T(OUT => "AASassetDB".PLC2Agent.Data.Initial_Time_Stamp);
   END_IF;
   #_w1 := "URI".Bits.Register[0] AND NOT #FlancoPos_Item_Completed;   // rising edge
   #FlancoPos_Item_Completed := "URI".Bits.Register[0];
   IF #_w1 THEN "Tag_4" := RD_LOC_T(OUT => "AASassetDB".PLC2Agent.Data.Final_Time_Stamp); END_IF;
END_REGION
END_ORGANIZATION_BLOCK

ORGANIZATION_BLOCK "Startup"   // OB100, STL, Startup
TITLE = "Complete Restart"
{ S7_Optimized_Access := 'TRUE' }
VERSION : 0.1
   VAR_INPUT
      LostRetentive : Bool;   // True if retentive data are lost
      LostRTC : Bool;   // True if date and time are lost
   END_VAR
BEGIN

REGION Network 1: Inicialización de las variables
         A     "MqttDB".control.connect;
         AN    "MqttDB".control.connect;
         =     "MqttDB".control.connect;

         A     "JSON_DeserializParamDB".execute;
         AN    "JSON_DeserializParamDB".execute;
         =     "JSON_DeserializParamDB".execute;